VERSION : 0.1
   STRUCT
      Offset_CP : Int;   // Offset cleaning piston
      Length_DrainPipe : Int;   // Length of drain pipe
      Diam_Piston : Int;   // Diameter piston
      ChokeSlot_min : Int;   // minimum choke slot at shot
      ChokeSlot_max : Int;   // maximum choke slot at shot
      RestTimeBack : S5Time;
      RestTimeFront : S5Time;
      RestTimeFrontManual : S5Time;
      IntervalCounts : Int;
      IntervalRestTimeBack : S5Time;
      IntervalRestTimeFront : S5Time;
      CP_after_PS : Bool;
      CP_withInterval : Bool;   // Cleaning piston with interval cleaning
      StepCleaningPiston : Bool;   // Equiped with a stepping cleaning piston
      ContrCleaningPiston : Bool;   // Equiped with a analog cleaning piston
      Spare_19 : Bool;
      Spare_20 : Bool;
      Spare_21 : Bool;
      Spare_22 : Bool;
      Spare_23 : Bool;
      Spare_24 : Bool;
      Spare_25 : Bool;
      Spare_26 : Bool;
      Spare_27 : Bool;
      Spare_28 : Bool;
      Spare_29 : Bool;
      Spare_30 : Bool;
   END_STRUCT;
END_TYPE

TYPE "UDT781_ParaPID_Ctrl"
TITLE = Parameters for PID Controller, used for pressure, temperature...
AUTHOR : KT242
VERSION : 0.1
   STRUCT
      ProportionalGain : Real;   // Reglerverstärkung
      ResetTime : Real;   // Integrationszeit
      DerivativeTime : Real;   // Differenzierzeit
      Spare12 : DWord;
   END_STRUCT;
END_TYPE

TYPE "UDT880_NozzleBypassO"
TITLE = Conf. ProCan Nozzle-Bypass-control overlapping
VERSION : 0.1
   STRUCT
      OverLBypassNozzle : Array[1..8] of Int;
      OverLNozzleBypass : Array[1..8] of Int;
   END_STRUCT;
   // OverLBypassNozzle[1] := 20;
   // OverLNozzleBypass[1] := 20;
END_TYPE

TYPE "UDT881_NozzleBypassD"
TITLE = Conf. ProCan Nozzle-Bypass-control delay
VERSION : 0.1
   STRUCT
      DelayShotStart : Array[1..8] of Int;
      DelayShotEnd : Array[1..8] of Int;
   END_STRUCT;
END_TYPE

TYPE "UDT886_ConfPos_Linearsen"
TITLE = Conf. ProCan position linear sensor piston
VERSION : 0.1
   STRUCT
      IniPos_oben : DInt := L#2000;   // Wert in Increments
      IniPos_unten : DInt := L#40000;   // Wert in Increments
   END_STRUCT;
END_TYPE

TYPE "UDT887_ConfLinerarsensor"
TITLE = Conf. ProCan linear sensor
VERSION : 0.1
   STRUCT
      Hersteller00 : Char := 'B';
      Hersteller01 : Char := 'A';
      Hersteller02 : Char := 'L';
      Hersteller03 : Char := 'L';
      Hersteller04 : Char := 'U';
      Hersteller05 : Char := 'F';
      Hersteller06 : Char := 'F';
      Hersteller07 : Char;
      GeraeteTyp00 : Char := 'B';
      GeraeteTyp01 : Char := 'T';
      GeraeteTyp02 : Char := 'L';
      GeraeteTyp03 : Char := '0';
      GeraeteTyp04 : Char := '2';
      GeraeteTyp05 : Char := '5';
      GeraeteTyp06 : Char := '0';
      GeraeteTyp07 : Char;
      SerienNrL : DWord := DW#16#12345678;
      SerienNrH : DWord;
      Aufloesung_Sensor : DInt := L#5000;
      Abtastrate : Int := 1;
   END_STRUCT;
END_TYPE

TYPE "UDT888_ConfAnaSPistonMH"
TITLE = Conf. ProCan analog steps cleaning piston
VERSION : 0.1
   STRUCT
      ConfAnaStepsPiston : Array[1..2] of "UDT899_ConfAnaStepPiston";
   END_STRUCT;
END_TYPE

TYPE "UDT895_ConfAnaCP_INI"
TITLE = Conf. ProCan input aproximate switch
VERSION : 0.1
   STRUCT
      CP_Home_DI_No_INI : Byte;   // Input number Ini Home position
      CP_Front_DI_No_INI : Byte;   // Input number Ini front position
   END_STRUCT;
END_TYPE

TYPE "UDT896_ConfAnaCP_Contr"
TITLE = Conf. ProCan controller cleaning piston
VERSION : 0.1
   STRUCT
      SettleTimeBeforeShot : Int := 100;
      CorrectionTimeatShot : Int := 100;
      RestTimeBack : Word;
      RestTimeFront : Word;
      TimeoutMovementForward : Word := W#16#1F4;   // 500 Hex
      TimeoutMovementBackward : Word := W#16#1F4;   // 500 Hex
      RearPosition : Int;
      CleaningPosition : Int := 1000;
      MaxPositionDuringShot : Int := 100;
      ContrSignals : Word;   // 1 means RestTimeFront starts when Piston is in front position
   END_STRUCT;
END_TYPE

TYPE "UDT897_ConfAnaContr"
TITLE = Conf. ProCan analog controller
VERSION : 0.1
   STRUCT
      LowValue : Int;   // low Value [as input calibration]
      HighValue : Int;   // high Value [as input calibration]
      ProportionalFactor : Int;   // proportional factor [0.01]
      IntegratorTime : Int;   // integrator time [ms]
      FilterTime : Int;   // filter time [ms]
      ModeFlags : Int;   // mode flags
      ZeroPointStep : Int;   // zero point step [as output calibration]
      NonLinearityPosition : Int;   // non-linearity position [as output calibration]
      NonLinearityStrength : Int;   // non-linearity strength [%]
      TolForControlloopOK : Int;   // tolerance for control loop ok bit
      TolBlockOfIntegrator : Int;
      MaxTimeBlockCalcIntegrat : Int;
   END_STRUCT;
END_TYPE

TYPE "UDT898_UserConfAnaCP"
VERSION : 0.1
   STRUCT
      MinThrottleGapDuringShot : Int;
      MaxThrottleGapDuringShot : Int;
      RearPosition : Int;
      CleaningPosition : Int;
      LengthExhaustingPipe : Int;
      RequestSetOffset : Bool;   // Request calculation of new offset for input position of cleaning pistonn
   END_STRUCT;
END_TYPE

TYPE "UDT899_ConfAnaStepPiston"
TITLE = Conf. ProCan analog steps cleaning piston
VERSION : 0.1
   STRUCT
      Options : Int;   // 1=Auto correction; 2=ignore approximation switch
      DurationStep0 : Int := 20;   // Duration step 0 [ms]
      DurationStep1 : Int := 20;   // Duration step 1 [ms]
      DurationStep2 : Int := 20;   // Duration step 2 [ms]
      DurationStep3 : Int := 20;   // Duration step 3 [ms]
      DurationStep4 : Int := 20;   // Duration step 4 [ms]
      VoltageStep0 : Int := 2000;   // Voltage step 0 [mV]
      VoltageStep1 : Int := 4000;   // Voltage step 1 [mV]
      VoltageStep2 : Int := 6000;   // Voltage step 2 [mV]
      VoltageStep3 : Int := 8000;   // Voltage step 3 [mV]
      VoltageStep4 : Int := 10000;   // Voltage step 4 [mV]
   END_STRUCT;
END_TYPE

TYPE "UDT900_ConfCalibFlow"
TITLE = Conf. PLC calibration flow value
VERSION : 0.1
   STRUCT
      Density : Int;
      Pulse_per_liter : Real;
      MaxFlow : Real;
      Factor : Real;
   END_STRUCT;
END_TYPE

TYPE "UDT901_ConfAna"
TITLE = Conf. ProCan analog value
VERSION : 0.1
   STRUCT
      Mode : Int := 2;   // mode
      Voltage_ZeroPos : Int;   // voltage [mV] for input value 0
      Value_10V : Word := W#16#2710;   // input value for 10 V or 138.5 W
      Time_Average_Value : Int := 200;   // time for moving average
   END_STRUCT;
END_TYPE

TYPE "UDT902_ConfFlow"
TITLE = Conf. ProCan flow value
VERSION : 0.1
   STRUCT
      Spare_2_0 : Bool;
      Spare_2_1 : Bool;
      Spare_2_2 : Bool;
      Spare_2_3 : Bool;
      Spare_2_4 : Bool;
      Spare_2_5 : Bool;
      Spare_2_6 : Bool;
      Spare_2_7 : Bool;
      single_phase : Bool;   // mode single phase flow input
      FPB_SPC0 : Bool;   // FPB pressure delivered by SPC 0
      FPB_SPC01 : Bool;   // FPB pressure delivered by SPC 1
      Pos_OUT : Bool;   // positive output if negative set value
      Spare_3_04 : Bool;
      Spare_3_05 : Bool;
      Spare_3_06 : Bool;
      Spare_3_07 : Bool;
      calibration : DInt := L#10000;   // calibration [0.0001 g/Imp]
      maximumflow : DInt := L#35000;   // maximum flow [0.01 g/s]
      controltime : Int := 200;   // closed loop control time [ms]
      controltime_FPB : Int := 500;   // closed loop control time [ms] during FPB
      time_average : Int := 200;   // time for moving average [ms]
      minimumVoltage : Int;   // minimum output voltage (-since 32768...+32767)
      maximumVoltage : Int := 32767;   // maximum output voltage (-32768...+32767)
      delayWarn_minVoltage : Int := 5000;   // time delay for warning bit of minimum voltage limit
      delayWarn_maxVoltage : Int := 5000;   // time delay for warning bit of maximum voltage limit
   END_STRUCT;
END_TYPE

TYPE "UDT903_ConfFlowTolQPU"
TITLE = Conf. ProCan quick pressure build up flow
VERSION : 0.1
   STRUCT
      flow_tolerance : DInt := L#1000;   // flow tolerance [0.01 g/s]
      timeout_for_FPB : Int := 5000;   // timeout for FPB [ms]
   END_STRUCT;
END_TYPE

TYPE "UDT904_ConfMHeadTimer"
TITLE = Conf. ProCan mixinghead timer
VERSION : 0.1
   STRUCT
      OpeningControlTime : Int := 500;   // opening control time [ms]
      ClosingControlTime : Int := 500;   // closing control time [ms]
      NozzleOpenDelay : Int;   // nozzle opening delay time [ms]
      NozzleClosingDelay : Int;   // nozzle closing delay time [ms]
      MH_ValveOutputNo : Int := 1;
      MH_ReleaseInputNo : Int;
      MH_APS_InputNo : Int := 9;
      NozzelOutputNo : Int;
   END_STRUCT;
END_TYPE

TYPE "UDT905_ConfTandemData"
VERSION : 0.1
   STRUCT
      start_pos_slowdown : DInt := L#10000;   // start position for slowdown
      start_pos_prep_change : DInt := L#80000;   // start position for preparing changeover
      P_value_start_vent : Int := 400;   // pressure value for start ventilating
      P_value_end_vent : Int := 100;   // pressure value for end ventilating
      allowed_pressure_tol : Int := 50;   // allowed pressure tolerance
      Set_pressure_diff : Int := -40;   // set pressure difference
      factor_filling_speed : Int := 200;   // factor for filling speed [0.01]
      factor_GDA_speed : Int := 100;   // factor for GDA speed [0.01]
      flow_filling_wo_circ : DInt := L#3000;   // flow for filling without circulation value [0.01 g/s]
      voltage_service_mode : Int := 1400;   // voltage for movement in service mode
      ignore_DPS_P_cross : Bool;   // .8 ignore DPS_PRESSURE_CROSS
      ignore_DPS_M_free : Bool;   // .9 ignore DPS_MOVE_FREE
      ignore_DPS_P_DEC : Bool;   // .10 DPS Pressure DEC auslassen
      Without_Aeration : Bool;   // .11 Without_Aeration
      spare_24_4 : Bool;   // .12
      spare_24_5 : Bool;   // .13
      spare_24_6 : Bool;   // .14
      spare_24_7 : Bool;   // .15
      idle_pos_at_bottom : Bool := TRUE;   // .0 idle position is at bottom
      aps_not_use_at_service : Bool;   // .1 approximate switch not use at service
      spare_25_2 : Bool;   // .2
      spare_25_3 : Bool;   // .3
      spare_25_4 : Bool;   // .4
      spare_25_5 : Bool;   // .5
      spare_25_6 : Bool;   // .6
      spare_25_7 : Bool;   // .7
      spare_26 : Int;
      spare_28 : Int;
   END_STRUCT;
END_TYPE

TYPE "UDT906_ConfTandemTimer"
VERSION : 0.1
   STRUCT
      tValve2Metering : Int;   // time between opening valves and start metering
      tControl : Int;   // time for delayed control after metering
      tMetering2Valve : Int;   // time between metering end and closing valves
      tValve2Ventilation : Int;   // time between closing valves and ventilation
      tVentilation : Int;   // maximum time for ventilation
      tValve2Filling : Int;   // time between opening valves and start filling
      tFilling2Valve : Int;   // time between filling end and closing valves
      tPauseFilling : Int;   // pause time after metering
      tValve2Buildup : Int;   // time between open valves and pressure build-up
      swapTime : Int;   // time for the ramp of swapover
      tmaxGDA : Int;   // max time of similar pressure build up
   END_STRUCT;
END_TYPE

TYPE "UDT907_ConfTandemState0"
VERSION : 0.1
   STRUCT
      DPS_NOT_ENABLED : Word;   // output mask for DPS_NOT_ENABLED
      not_used : Word;   // not_used
      DPS_START_METERING : Word;   // output mask for DPS_START_METERING
      DPS_METERING : Word;   // output mask for DPS_METERING
      DPS_RAMP_DOWN : Word;   // output mask for DPS_RAMP_DOWN
      DPS_DELAY_AFT_RMP : Word;   // output mask for DPS_DELAY_AFT_RMP
      DPS_DELAY_VALVE_C : Word;   // output mask for DPS_DELAY_VALVE_C
      DPS_PRESSURE_CROSS : Word;   // output mask for DPS_PRESSURE_CROSS
      DPS_PRESSURE_DEC : Word;   // output mask for DPS_PRESSURE_DEC
      DPS_DELAY_VENT_O : Word;   // output mask for DPS_DELAY_VENT_O
      DPS_VENTILATION : Word;   // output mask for DPS_VENTILATION
      DPS_WAIT_FOR_REFILL : Word;   // output mask for DPS_WAIT_FOR_REFILL
      DPS_DELAY_REFILL_O : Word;   // output mask for DPS_DELAY_REFILL_O
      DPS_REFILL : Word;   // output mask for DPS_REFILL
      DPS_DELAY_REFILL_C : Word;   // output mask for DPS_DELAY_REFILL_C
      DPS_DELAY_GDA : Word;   // output mask for DPS_DELAY_GDA
   END_STRUCT;
END_TYPE

TYPE "UDT908_ConfTandemState1"
VERSION : 0.1
   STRUCT
      DPS_MOVE_FREE : Word;   // output mask for DPS_MOVE_FREE
      DPS_WAIT_FOR_GDA : Word;   // output mask for DPS_WAIT_FOR_GDA
      DPS_START_METERING : Word;   // output mask for DPS_START_METERING
      DPS_GDA : Word;   // output mask for DPS_GDA
      DPS_READY_FOR_SWAP : Word;   // output mask for DPS_READY_FOR_SWAP
      DELAY_VALVE_O : Word;   // output mask for DPS_DELAY_VALVE_O
      DPS_RAMP_UP : Word;   // output mask for DPS_RAMP_UP
      not_used_14 : Word;
      not_used_16 : Word;
      DPS_SERVICE_WAIT : Word;   // output mask for DPS_SERVICE_WAIT
      DPS_SERVICE_DOWN : Word;   // output mask for DPS_SERVICE_DOWN
      DPS_SERVICE_UP : Word;   // output mask for DPS_SERVICE_UP
      not_used_24 : Word;
      DPS_SEARCH_REF : Word;   // output mask for DPS_SEARCH_REF
      not_used_28 : Word;
      not_used_30 : Word;
   END_STRUCT;
END_TYPE

TYPE "UDT909_ConfTandemStatef"
VERSION : 0.1
   STRUCT
      no_input_byte : Int;   // number of input byte (0...6)
      invert_mask_inputs : Word;   // invert mask for the inputs
      input_mask_upper_ini : Word;   // input mask for the upper initiator
      input_mask_lower_ini : Word;   // input mask for the lower initiator
   END_STRUCT;
END_TYPE

TYPE "UDT910_ProcessValue"
TITLE = Process value summary parameter
VERSION : 0.1
   STRUCT
      PV_SetV : "UDT911_PV_SetV";
      PV_ActV : "UDT916_Act_Prozess_Value";
      PV_Conf_ActV : "UDT912_PV_ActV_Conf";
   END_STRUCT;
END_TYPE

TYPE "UDT911_PV_SetV"
TITLE = Process Value set value, limits, limitcounter
VERSION : 0.1
   STRUCT
      Value : Real;   // Set value of the process value
      WarningLowerLimit : Real;   // Warning lower limit (setvalue - lower limit)
      WarningUpperLimit : Real;   // Warning upper limit (upper limit + setvalue)
      AlarmLowerLimit : Real;   // Alarm lower limit (setvalue - lower limit)
      AlarmUpperLimit : Real;   // Alarm upper limit (upper limit + setvalue)
   END_STRUCT;
END_TYPE

TYPE "UDT912_PV_ActV_Conf"
TITLE = Process value configuration actual value
VERSION : 0.1
   STRUCT
      ModulNo : Int;
      Address : Int;
      OffsetSignal : Int;   // Signal offset at zero point of measured value (axis intercept)
      Multiplier : Real;   // Multiplier to calculate actual value (gradient)
      MinValueSensor : Real;   // Min value of sensor
      MaxValueSensor : Real;   // Max value of sensor
      MaxSignalResolution : Real;   // Max. signal value from PLC or ProCan
   END_STRUCT;
END_TYPE

TYPE "UDT915_BuffResultSignal"
TITLE = State of shot result buffer
VERSION : 0.1
   STRUCT
      BufferReadPointer : Int;
      BufferWritePointer : Int := 1;
      BufferCounter : Int;
      Write : Bool;
      Read : Bool;
      Reset : Bool;
      WriteHFlag : Bool;
      ReadHFlag : Bool;
      ResetHFlag : Bool;
      BufferEmpty : Bool;
      BufferFull : Bool;
      NothingToRead : Bool;
      HF_BufferFullQuitt : Bool;
      HF_NewReadCycle : Bool;
      Spare73 : Bool;
      Spare74 : Bool;
      Spare75 : Bool;
      Spare76 : Bool;
      Spare77 : Bool;
      BufferLength : Int := 10;
      DB_No_Write : Int;   // Calculated DB number to write
      DB_No_Read : Int;
      DB_BufferLength : Int := 10;
      WarningLimitBuffer : Int;
      FaultBufferFull : Bool;
   END_STRUCT;
END_TYPE

TYPE "UDT916_Act_Prozess_Value"
TITLE = Process value actual value (min, max, average)
VERSION : 0.1
   STRUCT
      Value : Real;   // Actual value
      ValueState : Word;   // Bit0: Alarm low; Bit1: Warning low; Bit2: Warning overrunn; Bit3:Alarm overrun
   END_STRUCT;
END_TYPE

TYPE "UDT917_GenShotResult"
TITLE = Shot result general values (toolno.,shotno., ...)
VERSION : 0.1
   STRUCT
      SendData : Bool;   // Send Data to Shot Protocol
      ServiceShot : Bool;   // A Service shot was operated
      DateTime : Date_And_Time;
      RecipeNo : Int;
      RecipeID : DInt;
      ShotNo : Int;
      RobPrgNo : Int;
      Spare18 : Int;
      ToolNo : Int;
      ToolID : DInt;
      PartID : Int;
      CavityNo : Byte;
      SpareByte : Byte;
      StationNo : Byte;
      PlaceInStation : Byte;
      MH_No : Byte;
      Machine_No : Byte;
      ShotState : Array[0..15] of Bool;   // State 0 -> Error; State 1 -> Break; State 2 -> Service Shot
      MH_CompAlloc : Word;   // Components involved at shot
      ToolTemp : DInt;
      ToolPressure : DInt;
      PartWeight : Real;
      FoamingTime : Real;
      NitrogenValue_Inerting : Real;
      MH_OpeningTime : Real;   // Opening time of mixinghead [msec]
      MH_CloseingTime : Real;   // Closing time of mixinghead [msec]
      ToolStartTime : Date_And_Time;
      Toolname : String[10];
      Value_Nitrogen_Inerting : Real;
   END_STRUCT;
END_TYPE

TYPE "UDT918_CompShotResult"
TITLE = Shot result of the component values (flow, pressure ...)
VERSION : 0.1
   STRUCT
      Comp : Array[1..12] of "UDT940_FoamingResult";   // Foamingresults of the components involved at foaming
   END_STRUCT;
END_TYPE

TYPE "UDT919_ShotResult"
TITLE = Shot result summary
VERSION : 0.1
   STRUCT
      General : "UDT917_GenShotResult";
      Component : "UDT918_CompShotResult";
   END_STRUCT;
END_TYPE

TYPE "UDT920_Recipe"
TITLE = Production data recipe values
AUTHOR : KT242
VERSION : 0.1
   STRUCT
      ID_Recipe : DWord;   // Unique identifier of recipe
      CompTank : Array[1..12] of Struct   // Foaming data of component at tank 1-12
         WeightProportion : Int;   // Weight proportion of component at connected tank
         Pressure : Int;   // Pressure of component at connected tank 1/10 bar
         Spare1 : Int;
      END_STRUCT;
      Spare80 : Word;
   END_STRUCT;
END_TYPE

TYPE "UDT935_StatusShotSequenc"
TITLE = State shot sequence at a station
AUTHOR : KT242
VERSION : 0.1
   STRUCT
      Tool : "UDT930_Tool";
      StationNo : Byte;   // Stationumber of tool for foaming
      PartShot : Int;   // Part shot no. at faoming
      ToolNo : Int;   // Mixinghead number for next shot
      WorkCounter : DInt;   // Counts amount of tools foamed
      StartCycle : Bool;   // Start pulse for the foaming cycle
      StopCycle : Bool;   // Stop signal for foaming cycle
      StationActive : Bool;   // Work on this station is allready active
      ShotFound : Bool;   // bit that a shot for this machine was found
      StationFinished : Bool;   // Bit that all possible shots for this station have been checked
      Spare11_4 : Bool;
      Spare11_5 : Bool;
      Spare11_6 : Bool;
      Spare11_7 : Bool;
   END_STRUCT;
END_TYPE

TYPE "UDT940_FoamingResult"
VERSION : 0.1
   STRUCT
      "Name" : String[20];
      ComponentActive : Bool;
      MaterialConsumption : Real;   // Material consumption at shot
      Flow : Real;   // Flow of metering unit
      Flow_Set : Real;
      Pressure : Real;   // Pressure at metering unit
      Pressure_Set : Real;
      PressureMH : Real;   // Pressure at mixing head
      PressureMH_Set : Real;
      Temperature : Real;   // Temperature at filling tank
      Temperature_Set : Real;
      TemperatureMH : Real;   // Temperature at mixing head
      TemperatureMH_Set : Real;
      Mixingratio : Real;
      Mixingratio_Set : Real;
   END_STRUCT;
END_TYPE

TYPE "UDT940_FoamingResultLast10"
VERSION : 0.1
   STRUCT
      "Name" : String[20];
      StatusBitWarningFlow : Bool;
      StatusBitAlarmFlow : Bool;
      StatusBitWarningMixingratio : Bool;
      StatusBitAlarmMixingratio : Bool;
      StatusBitWarningPressure : Bool;
      StatusBitAlarmPressure : Bool;
      StatusBitWarningPressureMH : Bool;
      StatusBitAlarmPressureMH : Bool;
      StatusBitWarningTemperature : Bool;
      StatusBitAlarmTemperature : Bool;
      StatusBitWarningTemperatureMH : Bool;
      StatusBitAlarmTemperatureMH : Bool;
      StatusBitSpare14 : Bool;
      StatusBitSpare15 : Bool;
      StatusBitSpare16 : Bool;
      StatusBitSpare17 : Bool;
      Partcounter : Int;
      MaterialConsumption : Real;   // Material consumption at shot
      Flow : Real;   // Flow of metering unit
      Pressure : Real;   // Pressure at metering unit
      PressureMH : Real;   // Pressure at mixing head
      Temperature : Real;   // Temperature at filling tank
      TemperatureMH : Real;   // Temperature at mixing head
      Mixingratio : Real;
   END_STRUCT;
END_TYPE

TYPE "UDT1002_MH_Connection"
VERSION : 0.1
   STRUCT
      Pump_No : Int;   // Number of metering unit connected with mixing head
      Flow_HP_Circ : Real;   // Set value of flow at high pressure circulation
      Flow_red_Circ : Real;   // Set value of flow at reduced circulation
      Flow_LP_Circ : Real;   // Set value of flow at low pressure circulation
      Nozzel_delay_open : Real;
      Nozzel_delay_close : Real;
      FlowQPB : Real;   // Set value flow quick pressure build up [0.01 g/s]
      PressureQPB : Real;   // Set value pressure quick pressure build up
      HP_CircOverNozzle : Bool;   // high pressure recirculation over MH (not over bypass)
      Red_CircOverNozzle : Bool;   // reduced recirculation over MH (not over bypass)
      LP_CircOverNozzle : Bool;   // low pressure recirculation over MH (not over bypass)
      WithNozzle : Bool;   // Nozzle Control exist for these component
      HP_2Point_Flow : Bool;   // High pressure circulation with second speed
      Red_2Point_Flow : Bool;   // Reduced circulation with second speed
      LP_2Point_Flow : Bool;   // Low pressure circulation with second speed
      Exist : Bool;
      Spare08 : Bool;
      Spare09 : Bool;
      Spare10 : Bool;
      Spare11 : Bool;
      Spare12 : Bool;
      Spare13 : Bool;
      Spare14 : Bool;
      Spare15 : Bool;
      Spare27 : Byte;
   END_STRUCT;
END_TYPE

TYPE "UDT1003_MH_Connection_State"
VERSION : 0.1
   STRUCT
      "Name" : Array[1..6] of String[20];
      colour : Array[1..6] of Byte;
      MinFlow : Array[1..6] of Real;   // Maximun flow of pump [g/sec]
      MaxFlow : Array[1..6] of Real;   // Maximun flow of pump [g/sec]
      ActFlow : Array[1..6] of Real;   // Actual flow of pump [g/sec]
      HP_CircOverNozzle_Exist : Array[1..6] of Bool;
      Red_CircOverNozzle_Exist : Array[1..6] of Bool;
      LP_CircOverNozzle_Exist : Array[1..6] of Bool;
      HP_CircFlow_Exist : Array[1..6] of Bool;
      Red_CircFlow_Exist : Array[1..6] of Bool;
      LP_CircFlow_Exist : Array[1..6] of Bool;
      QPB_Exist : Array[1..6] of Bool;
      HP_2Point_Flow_Exist : Array[1..6] of Bool;   // High pressure circulation with second speed
      Red_2Point_Flow_Exist : Array[1..6] of Bool;   // Reduced circulation with second speed
      LP_2Point_Flow_Exist : Array[1..6] of Bool;   // Low pressure circulation with second speed
   END_STRUCT;
END_TYPE

TYPE "UDT1114_IF_Signals"
VERSION : 0.1
   STRUCT
      PrgNo : Byte;   // InputKM
      ExtP_OK : Bool;   // InputKM
      Strobe : Bool;   // InputKM
      Reserve1 : Bool;   // InputKM
      MH_open : Bool;   // InputKM
      CP_forward : Bool;   // InputKM
      Preparation : Bool;   // InputKM
      Start_Cleaning : Bool;   // InputKM
      Reserve3 : Bool;   // InputKM
      PU_OK : Bool;   // OutputKM
      Strobe_quitt : Bool;   // OutputKM
      cycle_run : Bool;   // OutputKM
      ready_for_shot : Bool;   // OutputKM
      shot_run : Bool;   // OutputKM
      shot_end : Bool;   // OutputKM
      Service_mode : Bool;   // OutputKM
      CP_is_forward : Bool;   // OutputKM
      Cleaning_finished : Bool;   // OutputKM
      Reserve31 : Bool;   // OutputKM
      Reserve32 : Bool;   // OutputKM
      Reserve33 : Bool;   // OutputKM
      Reserve34 : Bool;   // OutputKM
      Reserve35 : Bool;   // OutputKM
      Reserve36 : Bool;   // OutputKM
      Reserve37 : Bool;   // OutputKM
   END_STRUCT;
END_TYPE

TYPE "UDT1111_MouldCarrier"
VERSION : 0.1
   STRUCT
      Preparation : Bool;   // NonKM: Signal to start cycle
      StartFoaming : Bool;   // Non:KM: Signal to open mixinghead
      IN_Spare_01 : Bool;   // NonKM:
      IN_Spare_02 : Bool;   // NonKM:
      IN_Spare_03 : Bool;   // NonKM:
      IN_Spare_04 : Bool;   // NonKM:
      IN_Spare_05 : Bool;   // NonKM:
      IN_Spare_06 : Bool;   // NonKM:
      ShotEnds : Bool;   // KM: Signal shot ends
      Break : Bool;   // KM:Signal shot break // Fault
      OUT_Spare_01 : Bool;   // KM:
      OUT_Spare_02 : Bool;   // KM:
      OUT_Spare_03 : Bool;   // KM:
      OUT_Spare_04 : Bool;   // KM:
      OUT_Spare_05 : Bool;   // KM:
      OUT_Spare_06 : Bool;   // KM:
      NoFault : Bool;   // Status; No fault group 1 or 2 exist
      MachineAutomatic : Bool;   // Status: Machine in automatic mode
      MHAutomatic : Bool;   // Status: Mixinghead in automatic mode
      RobotAutomatic : Bool;   // Status: Robot in automatic mode
      WetShot : Bool;   // Status: Non service mode
      CycleRun : Bool;   // Status: Cycle runs
      ReadyForShot : Bool;   // Status: Ready for Shot
      ShotRun : Bool;   // Status: Shot run
      CPsisForward : Bool;   // Status: Cleaning pisteon is forward
      Status_Spare_01 : Bool;   // Status:
      Status_Spare_02 : Bool;   // Status:
      Status_Spare_03 : Bool;   // Status:
      Status_Spare_04 : Bool;   // Status:
      Status_Spare_05 : Bool;   // Status:
      Status_Spare_06 : Bool;   // Status:
      Status_Spare_07 : Bool;   // Status:
      ProgNumber : Bool;   // Status: Program number
      Fault_01 : Bool;   // Fault Message 01: Machine not in automatic mode
      Fault_02 : Bool;   // Fault Message 02: Mixinghead not in automatic mode
      Fault_03 : Bool;   // Fault Message 03: Robot not in automatik mode
      Fault_04 : Bool;   // Fault Message 04: Preparation signal interrupted
      Fault_05 : Bool;   // Fault Message 05: Enable signal not in time
      Fault_06 : Bool;   // Fault Message 06: Enable signal interrupted
      Fault_07 : Bool;   // Fault Message 07:
      Fault_08 : Bool;   // Fault Message 08:
   END_STRUCT;
END_TYPE

TYPE "UDT1112_APInterface"
VERSION : 0.1
   STRUCT
      PrgNo : Byte;   // nonKM:
      ExtP_OK : Bool;   // nonKM:
      Strobe : Bool;   // nonKM:
      StrobeInv : Bool;   // nonKM:
      MH_open : Bool;   // nonKM:
      CP_forward : Bool;   // nonKM:
      Preparation : Bool;   // nonKM:
      Start_Cleaning : Bool;   // nonKM:
      Stop : Bool;   // nonKM:
      PU_OK : Bool;   // KM:
      Strobe_quitt : Bool;   // KM:
      cycle_run : Bool;   // KM:
      ready_for_shot : Bool;   // KM:
      shot_run : Bool;   // KM:
      shot_end : Bool;   // KM:
      Service_mode : Bool;   // KM:
      CP_is_forward : Bool;   // KM:
      Cleaning_finished : Bool;   // KM:
      Reserve31 : Bool;   // KM:
      Reserve32 : Bool;   // KM:
      Reserve33 : Bool;   // KM:
      Reserve34 : Bool;   // KM:
      Reserve35 : Bool;   // KM:
      Reserve36 : Bool;   // KM:
      Reserve37 : Bool;   // KM:
      MachineAutomatic : Bool;   // Status: Machine in automatic mode
      MHAutomatic : Bool;   // Status: Mixinghead in automatic mode
      RobotAutomatic : Bool;   // Status: Robot in automatic mode
      WetShot : Bool;   // Status: Non service mode
      CycleRun : Bool;   // Status: Cycle runs
      ReadyForShot : Bool;   // Status: Ready for Shot
      ShotRun : Bool;   // Status: Shot run
      CPsisForward : Bool;   // Status: Cleaning pisteon is forward
      Status_Spare_01 : Bool;   // Status:
      Status_Spare_02 : Bool;   // Status:
      Status_Spare_03 : Bool;   // Status:
      Status_Spare_04 : Bool;   // Status:
      Status_Spare_05 : Bool;   // Status:
      Status_Spare_06 : Bool;   // Status:
      Status_Spare_07 : Bool;   // Status:
      Status_Spare_08 : Bool;   // Status:
      "Step" : Byte;   // Step number interface communication
      Fault_01 : Bool;   // Fault Message 01: Machine not in automatic mode
      Fault_02 : Bool;   // Fault Message 02: Mixinghead not in automatic mode
      Fault_03 : Bool;   // Fault Message 03: Robot not in automatik mode
      Fault_04 : Bool;   // Fault Message 04:
      Fault_05 : Bool;   // Fault Message 05:
      Fault_06 : Bool;   // Fault Message 06:
      Fault_07 : Bool;   // Fault Message 07:
      Fault_08 : Bool := false;   // Fault Message 08:
   END_STRUCT;
END_TYPE

TYPE "ABB_IRC5_Input"
VERSION : 0.0
   STRUCT
      diMotorOn : Bool;   // Systeminput: Switch ON the motors of the robot
      diMotorOff : Bool;   // Systeminput: Switch OFF the motors of the robot
      diStartProg : Bool;   // Systeminput: Start the robotprogram from the last position in the program
      diStartMain : Bool;   // Systeminput: Start the robotprogram from the beginning
      diStopProg : Bool;   // Systeminput: Stop the robotprogram
      diResetError : Bool;   // Systeminput: Reset an systemerror
      diResetEstop : Bool;   // Systeminput: Reset the emergencystop
      diQuickStop : Bool;   // Systeminput: Stop the robot directly and switch the break ON
      di_10_9 : Bool;   // Spare
      di_10_10 : Bool;   // Spare
      di_10_11 : Bool;   // Spare
      di_10_12 : Bool;   // Spare
      di_10_13 : Bool;   // Spare
      di_10_14 : Bool;   // Spare
      diBreak : Bool;   // Signal to call the interrupt 1
      diInterrupt : Bool;   // Signal to call the interrupt 2
      diStartCycle : Bool;   // Signal to start the robotcycle
      diReadProgNo : Bool;   // A programnumber can read from PLC
      diStartMoveMC : Bool;   // The robot can start with it´s movements
      diShotDigIn : Bool;   // The foaming enabling of the machine is existing
      diStartCleanMH : Bool;   // The robot can move to MH-Cleaningstation
      diCleanMHEnd : Bool;   // The MH-Cleaning is finished
      diStartBrushMH : Bool;   // Die Freigabe zum reinigen des MK's steht an (Bürstenstation ist bereit)
      diHomePrePos : Bool;   // Signal to move the robot from to the pre position
      diHomeToMaintP : Bool;   // Signal to move the robot from homeposition to maintenanceposition
      diMaintToHomeP : Bool;   // Signal to move the robot from maintenanceposition to homeposition
      diRobinSavepos : Bool;   // Signal das der Weg in die Grund/ Wartungsposition frei ist
      diProgBreak : Bool;   // Signal to break the program
      diJumpConveyer : Bool;   // Signal to jump the routine "Conveyer- Tracking"
      diStartSyncEPS : Bool;   // Signal to move the robot to the syncronisation switch
      diPLCWaitWobj : Bool;   // Signal to activate the waitwobj instruction
      diPLCDropWobj : Bool;   // Signal to drop the activ wobj
      diBackToRest : Bool;   // Signal to move the robot back to homeposition after foaming
      diHomeToMaint2 : Bool;   // Signal to move the robot from homeposition to maintenanceposition 2
      diStartEscape : Bool;   // Signal to move the robot to it´s escapeposition (anticollision)
      di10_36 : Bool;   // Spare
      di10_37 : Bool;   // Spare
      di10_38 : Bool;   // Spare
      di10_39 : Bool;   // Spare
      di10_40 : Bool;   // Spare
      di10_41 : Bool;   // Spare
      di10_42 : Bool;   // Spare
      di10_43 : Bool;   // Spare
      di10_44 : Bool;   // Reserve
      di10_45 : Bool;   // Reserve
      di10_46 : Bool;   // Reserve
      di10_47 : Bool;   // Reserve
      di10_48 : Bool;   // Reserve
      diAction_01 : Bool;   // Action 1 activ
      diAction_02 : Bool;   // Action 2 activ
      diAction_03 : Bool;   // Action 3 activ
      diAction_04 : Bool;   // Action 4 activ
      diAction_05 : Bool;   // Action 5 activ
      diAction_06 : Bool;   // Action 6 activ
      diAction_07 : Bool;   // Action 7 activ
      diAction_08 : Bool;   // Action 8 activ
      diAction_09 : Bool;   // Action 9 activ
      diAction_10 : Bool;   // Action 10 activ
      di10_59 : Bool;   // Spare
      di10_60 : Bool;   // Spare
      di10_61 : Bool;   // Spare
      di10_62 : Bool;   // Spare
      di10_63 : Bool;   // Spare
      di10_64 : Bool;   // Spare
      GIProgNo2 : Word;   // Programnumber 2 (right mould in mould carrier)
      giMouldCodeBit0 : Bool;   // Anzahl der Formen im Formträger (Gruppeingang Bit 0)
      giMouldCodeBit1 : Bool;   // Anzahl der Formen im Formträger (Gruppeingang Bit 1)
      di10_83 : Bool;   // Reserve
      di10_84 : Bool;   // Reserve
      di10_85 : Bool;   // Reserve
      di10_86 : Bool;   // Reserve
      di10_87 : Bool;   // Reserve
      di10_88 : Bool;   // Reserve
      GIMCNo : Byte;   // Nummer des Formträgers der Form// Abhängig vom MouldCode
      GIProgNo1 : Word;   // Programnumber 1 (left mould in mould carrier)
      GIShotTX1 : Word;   // Schußzeit des nächsten Teilschusses in 1/10 Sekunden
   END_STRUCT;
END_TYPE

TYPE "ABB_IRC5_Output"
VERSION : 0.0
   STRUCT
      doMotorOn : Bool;   // Systemoutput: Status for Motor OFF
      doMotorOff : Bool;   // Systemoutput: Status for Motor ON
      doCycleOn : Bool;   // Systemoutput: Robotprogram is running
      doIRBinAuto : Bool;   // Systemoutput: Robot is in operationmode AUTO
      doSysError : Bool;   // Systemoutput: Robot has an systemerror
      doEmStop_Akt : Bool;   // Systemoutput: Emergencystop at robot is active
      doMot_On_OK : Bool;   // Systemoutput: Automaticstopcicuites are OK
      doNullSpeed : Bool;   // Systemoutput: Conveyer is not moving
      doIRBInHome : Bool;   // Worldzoneoutput: Robot is in Homeposition
      doIRBInMaintP : Bool;   // Worldzoneoutput: Robot is in Maintenanceposition
      doIRBOutRange : Bool;   // Worldzoneoutput: Robot near the end of it´s workingarealimitation
      doIRBOutRangMC : Bool;   // Worldzoneoutput: Robot is out of the mould
      doIRBOutRanMC1 : Bool;   // Worldzoneoutput: Robot is outside the mould carrier 1
      doIRBOutRanMC2 : Bool;   // Worldzoneoutput: Robot is outside the mould carrier 2
      doIRBOutRanMC3 : Bool;   // Worldzoneoutput: Robot is outside the mould carrier 3
      doIRBOutRanMC4 : Bool;   // Worldzoneoutput: Robot is outside the mould carrier 4
      doCycleStarted : Bool;   // The programcycle is startet
      doCycleEnd : Bool;   // The programcycle is finished
      doProgNoReaded : Bool;   // The programnumber is readed
      doShotDigOut : Bool;   // 1st digital Shotware output // Signal to open the mixinghead
      doStopFormPLC : Bool;   // Signal to stop the foaming because the robotprogram has stoped
      doCloseMoulde : Bool;   // Signal that the robot is out of the mould
      doCleaningPLC : Bool;   // Control the mixinghead cleaner or a brush station
      doIRBSyncWobj : Bool;   // The robot is synchronized (Tracking)
      doRobWaitWobj : Bool;   // The robot is waiting for synchronizes (Tracking)
      doCleanOsziJet : Bool;   // Control the air for blow out the oszilation holes
      doBlowAir : Bool;   // Control the air for blow inside the mixinghead
      doCleanBrushOn : Bool;   // Control the cleaning for the mixinghead
      doShotDigOut2 : Bool;   // 2nd digital Shotware output
      doInPosTeach : Bool;   // The robot is in the position to teaching
      doConveyorStoped : Bool;   // The conveyor is stop
      doEpsControlPos : Bool;   // Signal to control the synchronization position
      doEpsSynchronized : Bool;   // Signal from Robot EPS is synchronize
      doEpsSyncSwitch : Bool;   // Signal from Robot sync switch is actuated
      doEpsSafeOut_1 : Bool;   // 1 Safe Output EPS
      doEpsSafeOut_2 : Bool;   // 2 Safe Output EPS
      doEpsSafeOut_3 : Bool;   // 3 Safe Output EPS
      doEpsSafeOut_4 : Bool;   // 4 Safe Output EPS
      doEpsSafeOut_5 : Bool;   // 5 Safe Output EPS
      doEpsPreWarn : Bool;   // Signal from pre warning robot sync
      doShotDigOut3 : Bool;   // 3rd digital Shotware output
      do01_042 : Bool;   // Reserve
      do10_43 : Bool;   // Reserve
      do10_44 : Bool;   // Reserve
      do10_45 : Bool;   // Reserve
      do10_46 : Bool;   // Reserve
      do10_47 : Bool;   // Reserve
      do10_48 : Bool;   // Reserve
      doAction_01 : Bool;   // Action 01 activ
      doAction_02 : Bool;   // Action 02 activ
      doAction_03 : Bool;   // Action 03 activ
      doAction_04 : Bool;   // Action 04 activ
      doAction_05 : Bool;   // Action 05 activ
      doAction_06 : Bool;   // Action 06 activ
      doAction_07 : Bool;   // Action 07 activ
      doAction_08 : Bool;   // Action 08 activ
      doAction_09 : Bool;   // Action 09 activ
      doAction_10 : Bool;   // Action 10 activ
      do10_59 : Bool;   // Reserve
      do10_60 : Bool;   // Reserve
      do10_61 : Bool;   // Reserve
      do10_62 : Bool;   // Reserve
      do10_63 : Bool;   // Reserve
      do10_64 : Bool;   // Reserve
      do10_65_80 : Word;   // Reserve
      do10_81_88 : Byte;   // Reserve
      goFormAktBit0 : Bool;   // Nummer der Form (1..3) welche zur Zeit bearbeitet wird (Gruppenausgang 0)
      goFormAktBit1 : Bool;   // Nummer der Form (1..3) welche zur Zeit bearbeitet wird (Gruppenausgang 1)
      go10_91 : Bool;   // Reserve
      go10_92 : Bool;   // Reserve
      go10_93 : Bool;   // Reserve
      go10_94 : Bool;   // Reserve
      go10_95 : Bool;   // Reserve
      go10_96 : Bool;   // Reserve
      GOError : Byte;   // Fehlernummer bei der Bearbeitung des Programms (Gruppenausgang)
      goxFIProgBit0 : Bool;   // Nummer des Faserprogrammes an den Rechner (Gruppenausgang der Shotware, Bit 0)
      goxFIProgBit1 : Bool;   // Nummer des Faserprogrammes an den Rechner (Gruppenausgang der Shotware, Bit 1)
      goxFIProgBit2 : Bool;   // Nummer des Faserprogrammes an den Rechner (Gruppenausgang der Shotware, Bit 2)
      goxFIProgBit3 : Bool;   // Nummer des Faserprogrammes an den Rechner (Gruppenausgang der Shotware, Bit 3)
      go10_117 : Bool;   // Reserve
      go10_118 : Bool;   // Reserve
      go10_119 : Bool;   // Reserve
      go10_120 : Bool;   // Reserve
      goOscixFIBit0 : Bool;   // Bit des Oszillierprogrammes // X1 (2'ter Gruppenausgang der Shotware, Bit 0)
      goOscixFIBit1 : Bool;   // Bit des Oszillierprogrammes // X2 (2'ter Gruppenausgang der Shotware, Bit 1)
      goOscixFIBit2 : Bool;   // Bit des Oszillierprogrammes // Y1 (2'ter Gruppenausgang der Shotware, Bit 2)
      goOscixFIBit3 : Bool;   // Bit des Oszillierprogrammes // Y2 (2'ter Gruppenausgang der Shotware, Bit 3)
      go10_125 : Bool;   // Reserve
      go10_126 : Bool;   // Reserve
      go10_127 : Bool;   // Reserve
      go10_128 : Bool;   // Reserve
   END_STRUCT;
END_TYPE

TYPE "ABB_IRC5_Messages"
VERSION : 0.0
   STRUCT
      Rob_ST_01_16 : Struct
         FLT_No_009 : Bool;
         FLT_No_010 : Bool;
         FLT_No_011 : Bool;
         FLT_No_012 : Bool;
         FLT_No_013 : Bool;
         FLT_No_014 : Bool;
         FLT_No_015 : Bool;
         FLT_No_016 : Bool;
         FLT_No_001 : Bool;
         FLT_No_002 : Bool;
         FLT_No_003 : Bool;
         FLT_No_004 : Bool;
         FLT_No_005 : Bool;
         FLT_No_006 : Bool;
         FLT_No_007 : Bool;
         FLT_No_008 : Bool;
      END_STRUCT;
      Rob_ST_17_32 : Struct
         FLT_No_025 : Bool;   // IRB auf dem Weg zur Form!
         FLT_No_026 : Bool;   // IRB wartet in der Vorposition der Form auf das Sartsignal der SPS!
         FLT_No_027 : Bool;   // IRB in Formträger <X> Formnummer <Y> Teilschuss <Z>
         FLT_No_028 : Bool;   // IRB außerhalb der Form nach dem Schäumen!
         FLT_No_029 : Bool;   // IRB auf dem Weg zum Reinigungsstation!
         FLT_No_030 : Bool;   // IRB ist in der Reinigungsstation! IRB wartet auf das Signal Reinigen starten
         FLT_No_031 : Bool;   // IRB ist in der Reinigungsstation! IRB wartet auf das Signal Reinigen beendet
         FLT_No_032 : Bool;   // IRB auf dem Weg zur Homeposition!
         FLT_No_017 : Bool;
         FLT_No_018 : Bool;
         FLT_No_019 : Bool;   // Falsche Programmnummer!
         FLT_No_020 : Bool;   // Es wurde seit 1h kein Startsignal an den Roboter übermittelt!
         FLT_No_021 : Bool;   // Das Signal <diReadProgNr> von der SPS zum IRB wird nicht zurückgesetzt!
         FLT_No_022 : Bool;   // Der von der SPS übertragene Mouldcode liegt außerhalb des zulässigen Bereiches
         FLT_No_023 : Bool;   // Der von der SPS übertragene Timecode liegt außerhalb des zulässigen Bereiches
         FLT_No_024 : Bool;   // Die aktuelle Schußzeit ist kleiner 1 sec!
      END_STRUCT;
      Rob_ST_33_48 : Struct
         FLT_No_041 : Bool;   // Bitte geben Sie die Formträger- nummer ein auf welcher die Form geteacht wird!
         FLT_No_042 : Bool;   // Starten Sie das Programm nun nur noch Schrittweise!
         FLT_No_043 : Bool;   // Zykluszeit 1 // Zykluszeit 2 // Zykluszeit 3 // Zykluszeit 4
         FLT_No_044 : Bool;   // Fehlerhafte Auswahl des FT! Es wurde kein Werkobjekt zugeordnet!
         FLT_No_045 : Bool;   // Programm wurde gestopt!
         FLT_No_046 : Bool;   // Soll das nächste Werkzeug optimiert werden?
         FLT_No_047 : Bool;   // Der Roboter wartet auf die Syncronisation!
         FLT_No_048 : Bool;   // Sprachauswahl!
         FLT_No_033 : Bool;   // IRB ist in der Homeposition!
         FLT_No_034 : Bool;   // IRB auf dem Weg zur Wartungsposition!
         FLT_No_035 : Bool;   // IRB ist in der Wartungsposition!
         FLT_No_036 : Bool;   // IRB wartet auf <Zyklus-Start> Signal!
         FLT_No_037 : Bool;   // IRB liest Daten von der SPS!
         FLT_No_038 : Bool;   // IRB wartet auf <Schäumen-Start> Signal von der SPS!
         FLT_No_039 : Bool;   // IRB wartet auf <Schäumen-Beenden> Signal von der SPS!
         FLT_No_040 : Bool;   // Bitte geben Sie das zu teachende Programm ein!
      END_STRUCT;
      Rob_ST_49_64 : Struct
         FLT_No_057 : Bool;   // Angewähle Optionen: Shotware: Ja // Tracking : No // Programm Verschiebung: No
         FLT_No_058 : Bool;   // Angewähle Optionen: Shotware: No // Tracking : Ja // Programm Verschiebung: Ja
         FLT_No_059 : Bool;   // Angewähle Optionen: Shotware: No // Tracking : Ja // Programm Verschiebung: No
         FLT_No_060 : Bool;   // Angewähle Optionen: Shotware: No // Tracking : No // Programm Verschiebung: Ja
         FLT_No_061 : Bool;   // Angewähle Optionen: Shotware: No // Tracking : No // Programm Verschiebung: No
         FLT_No_062 : Bool;   // Zum Ändern der Daten benötigen Sie ein Password! Möchten Sie diese Daten ändern
         FLT_No_063 : Bool;   // Bitte geben Sie das Password ein. Password:
         FLT_No_064 : Bool;   // Sie sind nicht berechtigt diese Daten zu ändern!
         FLT_No_049 : Bool;   // Sprachauswahl!
         FLT_No_050 : Bool;   // Sollen die Texte auf dem Bildschirm angezeigt werden?
         FLT_No_051 : Bool;   // Wurde der Roboter mit der Option <SHOTWARE> gebooted?
         FLT_No_052 : Bool;   // Wurde der Roboter mit der Option <Conveyer - Tracking> gebooted?
         FLT_No_053 : Bool;   // Soll das Bewegugsprogram auf einem Formträger verschoben werden?
         FLT_No_054 : Bool;   // Angewähle Optionen: Shotware: Ja // Tracking : Ja // Programm Verschiebung: Ja
         FLT_No_055 : Bool;   // Angewähle Optionen: Shotware: Ja // Tracking : Ja // Programm Verschiebung: No
         FLT_No_056 : Bool;   // Angewähle Optionen: Shotware: Ja // Tracking : No // Programm Verschiebung: Ja
      END_STRUCT;
      Rob_ST_65_80 : Struct
         FLT_No_073 : Bool;
         FLT_No_074 : Bool;
         FLT_No_075 : Bool;
         FLT_No_076 : Bool;
         FLT_No_077 : Bool;
         FLT_No_078 : Bool;
         FLT_No_079 : Bool;
         FLT_No_080 : Bool;
         FLT_No_065 : Bool;   // Geschwindigkeits - Override <100% !!! Soll dieser nun auf 100% gesetzt werden?
         FLT_No_066 : Bool;   // KM-SOFTWARE!!! SIE sind nicht Autorisiert diese Software zu benutzen!
         FLT_No_067 : Bool;   // Bewegungszeit 1 // Bewegungszeit 2 // Bewegungszeit 3 // Bewegungszeit 4
         FLT_No_068 : Bool;   // Starten Sie nun das zu teachende Programm über das Menü Spezial - 4!
         FLT_No_069 : Bool;   // Abbruch Datenlesen von der SPS!
         FLT_No_070 : Bool;
         FLT_No_071 : Bool;
         FLT_No_072 : Bool;
      END_STRUCT;
   END_STRUCT;
END_TYPE

TYPE "UDT1201_ProCanAddress"
VERSION : 0.1
   STRUCT
      Input : "UDT1210_ProCan_Input";
      Output : "UDT1220_ProCan_Output";
      Address : "UDT1230_ProCanUnitNo";
      Flag_Modul_OK : Bool;
      Flag_Modul_NOK : Bool;   // _
      Spare_02 : Bool;
      Spare_03 : Bool;
      Spare_04 : Bool;
      Spare_05 : Bool;
      Spare_06 : Bool;
      Spare_07 : Bool;
      Spare_08 : Bool;
      Spare_09 : Bool;
      Spare_010 : Bool;
      Spare_011 : Bool;
      Spare_012 : Bool;
      Spare_013 : Bool;
      Spare_014 : Bool;
      Spare_015 : Bool;
   END_STRUCT;
END_TYPE

TYPE "UDT1210_ProCan_Input"
VERSION : 0.1
   STRUCT
      Telegram : Int;
      Telegram_Reserve : Int;
   END_STRUCT;
END_TYPE

TYPE "UDT1220_ProCan_Output"
VERSION : 0.1
   STRUCT
      Reserve01 : Int;
      Telegram_Recive : Int;   // Address recive telegram data (36 byte)
   END_STRUCT;
END_TYPE

TYPE "UDT1230_ProCanUnitNo"
VERSION : 0.1
   STRUCT
      MachineNo : Int;
      FlowNo01 : Int;
      FlowNo02 : Int;
      FlowNo03 : Int;
      FlowNo04 : Int;
      MixingheadNo01 : Int;
      MixingheadNo02 : Int;
      BypassNozzelNo01 : Int;
      BypassNozzelNo02 : Int;
      MeteringPistonNo01 : Int;
      MeteringPistonNo02 : Int;
      MeteringPistonNo03 : Int;
      MeteringPistonNo04 : Int;
      TandemNo01 : Int;
      TandemNo02 : Int;
      PLC_No01 : Int;
      PLC_No02 : Int;
      PLC_No03 : Int;
      PLC_No04 : Int;
   END_STRUCT;
END_TYPE

TYPE "UDT1232_ProCanIO_MH"
VERSION : 0.1
   STRUCT
      Ref_Digital_Input : Int;
      Ref_MH_ShotTime : Int;
      Ref_MH_Opening_Time : Int;
      Ref_MH_Closing_Time : Int;
      Ref_MH_State : Int;
      Ref_PLC_State : Int;
      Ref_CP_State : Int;
      Ref_Digital_Output : Int;
      Ref_ShotTimeSetValue : Int;
      Ref_ServiceProduction : Int;
      Ref_MixingheadControl : Int;
      Ref_PLC_comand_SP : Int;   // Address Command word cLose loop control steering piston
      Ref_PLC_comand_CP : Int;   // Address Command word cLose loop control cleaning piston
      Ref_PLC_set_value_SP : Int;   // Address set value cLose loop control steering piston
      Ref_PLC_set_value_CP : Int;   // Address set value cLose loop control cleaning piston
      Ref_NozzelBypassControl : Int;   // Address bypass control (byte)
      Ref_NozzelBypassSetOut : Int;   // Address set nozzels of bypass (byte)
      Ref_Reserve : Int;
      Ref_OK : Bool;
      MH_Channel_01 : Bool;
      MH_Channel_02 : Bool;
      Spare_03 : Bool;
      Spare_04 : Bool;
      Spare_05 : Bool;
      Spare_06 : Bool;
      Spare_07 : Bool;
   END_STRUCT;
END_TYPE

TYPE "UDT1233_ProCanIO_Flow"
VERSION : 0.1
   STRUCT
      Ref_Act_FlowValue : Int;
      Ref_Act_FlowState : Int;
      Ref_Set_FlowRate : Int;
      Ref_Set_FlowRateQPB : Int;
      Ref_Act_PressureQPB : Int;
      Ref_Set_SWO_PressureQPB : Int;
      Ref_Set_FlowIndexFlags : Int;
      Ref_TandemStatus : Int;
      Ref_TandemComand : Int;
      Ref_PistonPosition : Int;
      Ref_OK : Bool;
   END_STRUCT;
END_TYPE

TYPE "UDT1440_BuffProCan"
VERSION : 0.1
   STRUCT
      muxin : Bool;   // Toggelbit an dem Rechner das sich die Sendedaten geändert haben
      muxout : Bool;   // Toggelbit von dem Rechner das die Sendedatenänderung erkannt wurde
      ProCanMessage : Bool;   // Wird benötigt wenn Sendedaten mit dem ProCan- Modul ausgetauscht werden sollen
      ProCanBufferEmpty : Bool;   // Der Empfangsdatenbereich zum ProCan- Modul ist leer, bereit zum neuen Transfer
      transferBufferEmpty : Bool;   // Der Empfangsdatenbereich zur Steuerung ist leer, bereit zum neuen Transfer
      Spare_0_5 : Bool;   // Reserve in der Verwaltung des Empfangsbereiches
      Spare_0_6 : Bool;   // Reserve in der Verwaltung des Empfangsbereiches
      Spare_0_7 : Bool;   // Reserve in der Verwaltung des Empfangsbereiches
      Length : Byte;   // Länge der aktuell übertragenen Empfangsdaten (Max. 32 Byte)
      ID : Byte;   // Kennung der aktuellen Empfangsdaten zur Unterscheidung was empfangen wurde
      ID2 : Byte;   // 2. Kennung der aktuellen Empfangsdaten zur Unterscheidung des Blockes
      Data : "UDT1441_BuffProCanData";
   END_STRUCT;
END_TYPE

TYPE "UDT1441_BuffProCanData"
VERSION : 0.1
   STRUCT
      Data_01_04 : DWord;   // Send buffer Bytes 01- 04
      Data_05_08 : DWord;   // Send buffer Bytes 05- 08
      Data_09_12 : DWord;   // Send buffer Bytes 09- 12
      Data_13_16 : DWord;   // Send buffer Bytes 13- 16
      Data_17_20 : DWord;   // Send buffer Bytes 17- 20
      Data_21_24 : DWord;   // Send buffer Bytes 21- 24
      Data_25_28 : DWord;   // Send buffer Bytes 25- 28
      Data_29_32 : DWord;   // Send buffer Bytes 29- 32
   END_STRUCT;
END_TYPE

TYPE "UDT1442_BufferTrans"
VERSION : 0.1
   STRUCT
      ID_Data_sending : Byte;
      ID2_Data_sending : Byte;
      ID_Mask_sending : Byte;
      No_TransferedBlocks : Byte;
   END_STRUCT;
END_TYPE

